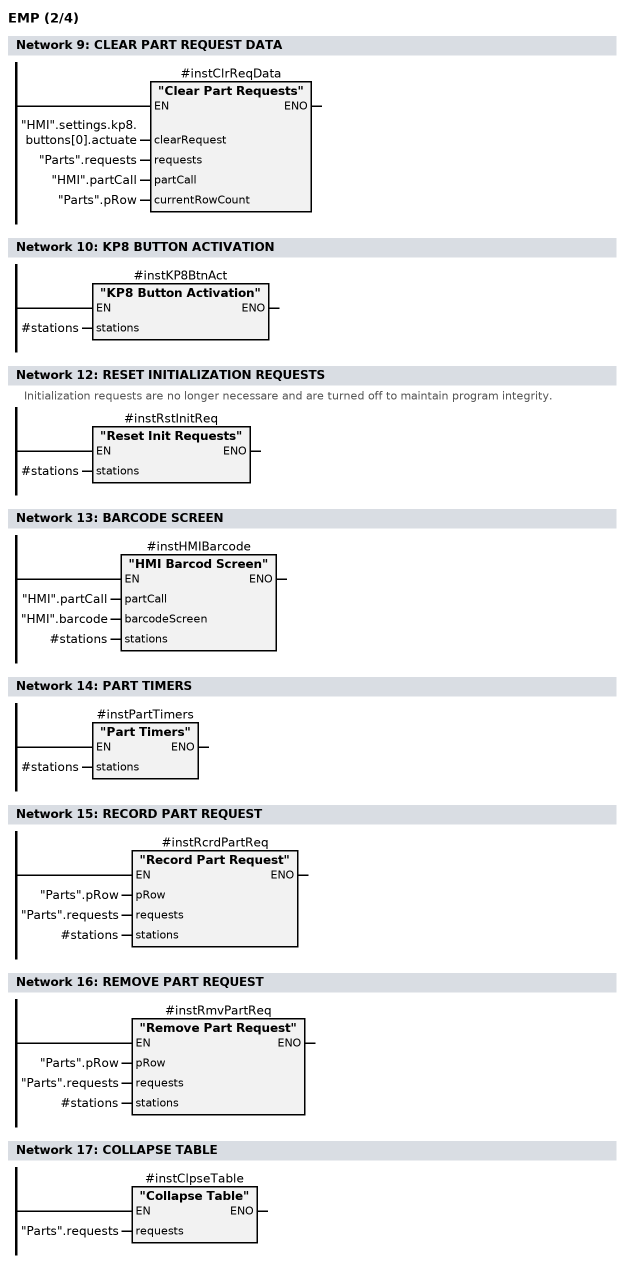
   RUNG wire#powerrail
      #instClrReqData(clearRequest := "HMI".settings.kp8.buttons[0].actuate, requests := "Parts".requests, partCall := "HMI".partCall, currentRowCount := "Parts".pRow)
   END_RUNG
   // the same network as SCL:
   #instClrReqData(clearRequest := "HMI".settings.kp8.buttons[0].actuate,   // "Clear Part Requests"
                   requests := "Parts".requests,
                   partCall := "HMI".partCall,
                   currentRowCount := "Parts".pRow);
END_REGION

REGION Network 10: KP8 BUTTON ACTIVATION
   RUNG wire#powerrail
      #instKP8BtnAct(stations := #stations)
   END_RUNG
   // the same network as SCL:
   #instKP8BtnAct(stations := #stations);   // "KP8 Button Activation"
END_REGION

REGION Network 11 (SCL): KP8 DRIVER CALLS
   REGION "LOOP THROUGH STATIONS"
       FOR #i := 0 TO "stnCount" DO
           #instKP8Drvs[#i](btnIn := #stations.me[#i].kp8In,
                            hardInit := #stations.me[#i].init.hard,
                            softInit := #stations.me[#i].init.soft,
                            btn0Activate := #stations.me[#i].kp8Config.activate[0],
                            btn0Mode := #stations.me[#i].kp8Config.mode[0],
                            btn0Group := #stations.me[#i].kp8Config.group[0],
                            btn0Flash := #stations.me[#i].kp8Config.flash[0],
                            btn0ColorOn1 := #stations.me[#i].kp8Config.colorOn1[0],
                            btn0ColorOn2 := #stations.me[#i].kp8Config.colorOn2[0],
                            btn0ColorOff := #stations.me[#i].kp8Config.colorOff[0],
                            btn1Activate := #stations.me[#i].kp8Config.activate[1],
                            btn1Mode := #stations.me[#i].kp8Config.mode[1],
                            btn1Group := #stations.me[#i].kp8Config.group[1],
                            btn1Flash := #stations.me[#i].kp8Config.flash[1],
                            btn1ColorOn1 := #stations.me[#i].kp8Config.colorOn1[1],
                            btn1ColorOn2 := #stations.me[#i].kp8Config.colorOn2[1],
                            btn1ColorOff := #stations.me[#i].kp8Config.colorOff[1],
                            btn2Activate := #stations.me[#i].kp8Config.activate[2],
                            btn2Mode := #stations.me[#i].kp8Config.mode[2],
                            btn2Group := #stations.me[#i].kp8Config.group[2],
                            btn2Flash := #stations.me[#i].kp8Config.flash[2],
                            btn2ColorOn1 := #stations.me[#i].kp8Config.colorOn1[2],
                            btn2ColorOn2 := #stations.me[#i].kp8Config.colorOn2[2],
                            btn2ColorOff := #stations.me[#i].kp8Config.colorOff[2],
                            btn3Activate := #stations.me[#i].kp8Config.activate[3],
                            btn3Mode := #stations.me[#i].kp8Config.mode[3],
                            btn3Group := #stations.me[#i].kp8Config.group[3],
                            btn3Flash := #stations.me[#i].kp8Config.flash[3],
                            btn3ColorOn1 := #stations.me[#i].kp8Config.colorOn1[3],
                            btn3ColorOn2 := #stations.me[#i].kp8Config.colorOn2[3],
                            btn3ColorOff := #stations.me[#i].kp8Config.colorOff[3],
                            btn4Activate := #stations.me[#i].kp8Config.activate[4],
                            btn4Mode := #stations.me[#i].kp8Config.mode[4],
                            btn4Group := #stations.me[#i].kp8Config.group[4],
                            btn4Flash := #stations.me[#i].kp8Config.flash[4],
                            btn4ColorOn1 := #stations.me[#i].kp8Config.colorOn1[4],
                            btn4ColorOn2 := #stations.me[#i].kp8Config.colorOn2[4],
                            btn4ColorOff := #stations.me[#i].kp8Config.colorOff[4],
                            btn5Activate := #stations.me[#i].kp8Config.activate[5],
                            btn5Mode := #stations.me[#i].kp8Config.mode[5],
                            btn5Group := #stations.me[#i].kp8Config.group[5],
                            btn5Flash := #stations.me[#i].kp8Config.flash[5],
                            btn5ColorOn1 := #stations.me[#i].kp8Config.colorOn1[5],
                            btn5ColorOn2 := #stations.me[#i].kp8Config.colorOn2[5],
                            btn5ColorOff := #stations.me[#i].kp8Config.colorOff[5],
                            btn6Activate := #stations.me[#i].kp8Config.activate[6],
                            btn6Mode := #stations.me[#i].kp8Config.mode[6],
                            btn6Group := #stations.me[#i].kp8Config.group[6],
                            btn6Flash := #stations.me[#i].kp8Config.flash[6],
                            btn6ColorOn1 := #stations.me[#i].kp8Config.colorOn1[6],
                            btn6ColorOn2 := #stations.me[#i].kp8Config.colorOn2[6],
                            btn6ColorOff := #stations.me[#i].kp8Config.colorOff[6],
                            btn7Activate := #stations.me[#i].kp8Config.activate[7],
                            btn7Mode := #stations.me[#i].kp8Config.mode[7],
                            btn7Group := #stations.me[#i].kp8Config.group[7],
                            btn7Flash := #stations.me[#i].kp8Config.flash[7],
                            btn7ColorOn1 := #stations.me[#i].kp8Config.colorOn1[7],
                            btn7ColorOn2 := #stations.me[#i].kp8Config.colorOn2[7],
                            btn7ColorOff := #stations.me[#i].kp8Config.colorOff[7],
                            btnStatesOut => #stations.me[#i].btnStates,
                            btnColorsOut => #stations.me[#i].kp8Out);
       END_FOR;
   END_REGION
END_REGION

REGION Network 12: RESET INITIALIZATION REQUESTS
   // Initialization requests are no longer necessare and are turned off to maintain program integrity.
   RUNG wire#powerrail
      #instRstInitReq(stations := #stations)
   END_RUNG
   // the same network as SCL:
   #instRstInitReq(stations := #stations);   // "Reset Init Requests"
END_REGION

REGION Network 13: BARCODE SCREEN
   RUNG wire#powerrail
      #instHMIBarcode(partCall := "HMI".partCall, barcodeScreen := "HMI".barcode, stations := #stations)
   END_RUNG
   // the same network as SCL:
   #instHMIBarcode(partCall := "HMI".partCall, barcodeScreen := "HMI".barcode, stations := #stations);   // "HMI Barcod Screen"
END_REGION

REGION Network 14: PART TIMERS
   RUNG wire#powerrail
      #instPartTimers(stations := #stations)
   END_RUNG
   // the same network as SCL:
   #instPartTimers(stations := #stations);   // "Part Timers"
END_REGION

REGION Network 15: RECORD PART REQUEST
   RUNG wire#powerrail
      #instRcrdPartReq(pRow := "Parts".pRow, requests := "Parts".requests, stations := #stations)
   END_RUNG
   // the same network as SCL:
   #instRcrdPartReq(pRow := "Parts".pRow, requests := "Parts".requests, stations := #stations);   // "Record Part Request"
END_REGION

REGION Network 16: REMOVE PART REQUEST
   RUNG wire#powerrail
      #instRmvPartReq(pRow := "Parts".pRow, requests := "Parts".requests, stations := #stations)
   END_RUNG
   // the same network as SCL:
   #instRmvPartReq(pRow := "Parts".pRow, requests := "Parts".requests, stations := #stations);   // "Remove Part Request"
END_REGION

REGION Network 17: COLLAPSE TABLE
   RUNG wire#powerrail
      #instClpseTable(requests := "Parts".requests)
   END_RUNG
   // the same network as SCL:
   #instClpseTable(requests := "Parts".requests);   // "Collapse Table"
END_REGION

REGION Network 18: LOG REQUESTS
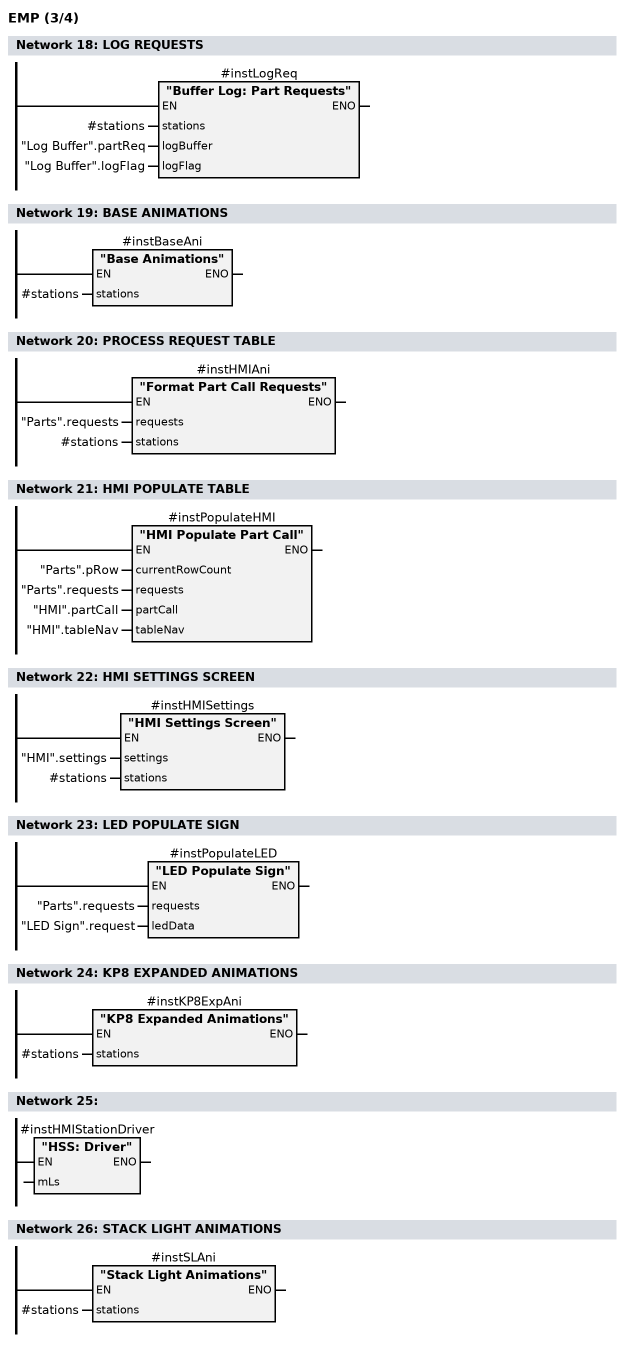
   RUNG wire#powerrail
      #instLogReq(stations := #stations, logBuffer := "Log Buffer".partReq, logFlag := "Log Buffer".logFlag)
   END_RUNG
   // the same network as SCL:
   #instLogReq(stations := #stations, logBuffer := "Log Buffer".partReq, logFlag := "Log Buffer".logFlag);   // "Buffer Log: Part Requests"
END_REGION

REGION Network 19: BASE ANIMATIONS
   RUNG wire#powerrail
      #instBaseAni(stations := #stations)
   END_RUNG
   // the same network as SCL:
   #instBaseAni(stations := #stations);   // "Base Animations"
END_REGION

REGION Network 20: PROCESS REQUEST TABLE
   RUNG wire#powerrail
      #instHMIAni(requests := "Parts".requests, stations := #stations)
   END_RUNG
   // the same network as SCL:
   #instHMIAni(requests := "Parts".requests, stations := #stations);   // "Format Part Call Requests"
END_REGION

REGION Network 21: HMI POPULATE TABLE
   RUNG wire#powerrail
      #instPopulateHMI(currentRowCount := "Parts".pRow, requests := "Parts".requests, partCall := "HMI".partCall, tableNav := "HMI".tableNav)
   END_RUNG
   // the same network as SCL:
   #instPopulateHMI(currentRowCount := "Parts".pRow,   // "HMI Populate Part Call"
                    requests := "Parts".requests,
                    partCall := "HMI".partCall,
                    tableNav := "HMI".tableNav);
END_REGION

REGION Network 22: HMI SETTINGS SCREEN
   RUNG wire#powerrail
      #instHMISettings(settings := "HMI".settings, stations := #stations)
   END_RUNG
   // the same network as SCL:
   #instHMISettings(settings := "HMI".settings, stations := #stations);   // "HMI Settings Screen"
END_REGION

REGION Network 23: LED POPULATE SIGN
   RUNG wire#powerrail
      #instPopulateLED(requests := "Parts".requests, ledData := "LED Sign".request)
   END_RUNG
   // the same network as SCL:
   #instPopulateLED(requests := "Parts".requests, ledData := "LED Sign".request);   // "LED Populate Sign"
END_REGION

REGION Network 24: KP8 EXPANDED ANIMATIONS
   RUNG wire#powerrail
      #instKP8ExpAni(stations := #stations)
   END_RUNG
   // the same network as SCL:
   #instKP8ExpAni(stations := #stations);   // "KP8 Expanded Animations"
END_REGION

REGION Network 25
   RUNG wire#powerrail
      #instHMIStationDriver(mLs :=)
   END_RUNG
   // the same network as SCL:
   #instHMIStationDriver();   // "HSS: Driver"
END_REGION

REGION Network 26: STACK LIGHT ANIMATIONS
   RUNG wire#powerrail
      #instSLAni(stations := #stations)
   END_RUNG
   // the same network as SCL:
   #instSLAni(stations := #stations);   // "Stack Light Animations"
END_REGION

REGION Network 27: GLOBAL TO SIMULATION
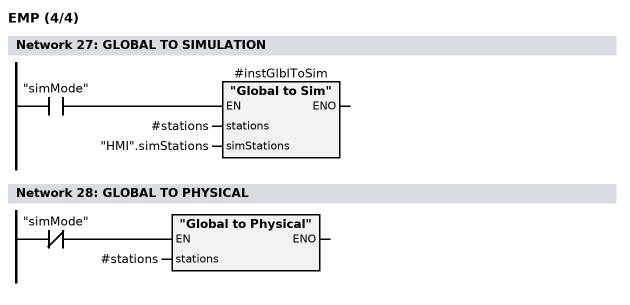
   RUNG wire#powerrail
      Contact( "simMode" )
      #instGlblToSim(stations := #stations, simStations := "HMI".simStations)
   END_RUNG
   // the same network as SCL:
   IF "simMode" THEN
       #instGlblToSim(stations := #stations, simStations := "HMI".simStations);   // "Global to Sim"
   END_IF;
END_REGION

REGION Network 28: GLOBAL TO PHYSICAL
   RUNG wire#powerrail
      I_Contact( "simMode" )
      "Global to Physical"(stations := #stations)
   END_RUNG
   // the same network as SCL:
   IF NOT "simMode" THEN "Global to Physical"(stations := #stations); END_IF;
END_REGION
END_FUNCTION_BLOCK

// folder: HMI Select Station

FUNCTION_BLOCK "HSS: Driver"   // FB32, LAD
{ S7_Optimized_Access := 'TRUE' }
VERSION : 0.1
   VAR_INPUT
      mLs : "Menu: Libraries";
   END_VAR
   VAR
      recipeSelector : Int;
      r1 : DInt;
      instHSSMenuSelection : "HSS: Menu Selection";
   END_VAR
   VAR_TEMP
      i : Int;
   END_VAR
BEGIN

REGION Network 1
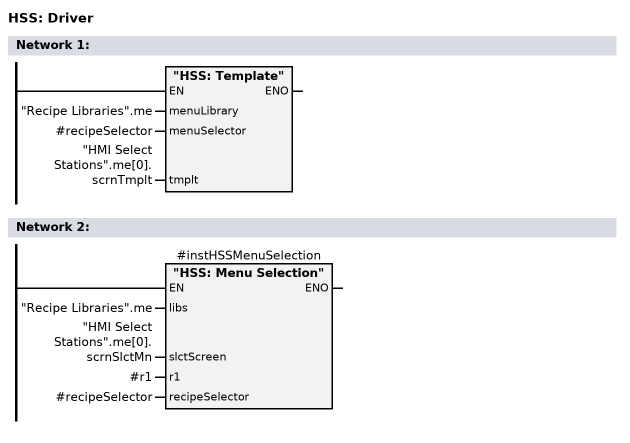
   RUNG wire#powerrail
      "HSS: Template"(menuLibrary := "Recipe Libraries".me, menuSelector := #recipeSelector, tmplt := "HMI Select Stations".me[0].scrnTmplt)
   END_RUNG
   // the same network as SCL:
   "HSS: Template"(menuLibrary := "Recipe Libraries".me,
                   menuSelector := #recipeSelector,
                   tmplt := "HMI Select Stations".me[0].scrnTmplt);
END_REGION

REGION Network 2
   RUNG wire#powerrail
      #instHSSMenuSelection(libs := "Recipe Libraries".me, slctScreen := "HMI Select Stations".me[0].scrnSlctMn, r1 := #r1, recipeSelector := #recipeSelector)
   END_RUNG
   // the same network as SCL:
   #instHSSMenuSelection(libs := "Recipe Libraries".me,   // "HSS: Menu Selection"
                         slctScreen := "HMI Select Stations".me[0].scrnSlctMn,
                         r1 := #r1,
                         recipeSelector := #recipeSelector);
END_REGION
END_FUNCTION_BLOCK

FUNCTION_BLOCK "HSS: Part Selection"   // FB33, SCL
{ S7_Optimized_Access := 'TRUE' }
VERSION : 0.1
BEGIN
END_FUNCTION_BLOCK

FUNCTION_BLOCK "HSS: Menu Selection"   // FB35, SCL
{ S7_Optimized_Access := 'TRUE' }
VERSION : 0.1
   VAR_INPUT
      libs : "Menu: Libraries";
   END_VAR
   VAR_IN_OUT
      slctScreen : "HSS: Menu Selection Screen";
      r1 : DInt;
      recipeSelector : Int;
   END_VAR
   VAR
      old : Struct
         navPress : Bool;
      END_STRUCT;
      instTableNavigation : "Table Navigatio";
   END_VAR
   VAR_TEMP
      eval : "HSS: Menu Selection Screen";
      pbs : Array[0..#pbFlagCnt] of Bool;
      POS : DInt;
      status : DInt;
      i : Int;
      btnNum : Int;
      pRowVisLbl : Int;
      pRowInvisLbl : Int;
      pRecipeInvisLbl : Int;
      pRecipeVisLbl : Int;
      pRecipeLib : Int;
      pRowTxt : Int;
      pRecipeTxt : Int;
      shifter : DWord;
      btnsAsBool : Array[0..31] of Bool;
      rows : Array[0..99] of DInt;
      offset : DInt;
      navPress : Bool;
      selPress : Bool;
      maxRows : DInt;
   END_VAR
   VAR CONSTANT
      pbFlagCnt : Int := 31;
      btnCnt : Int := 5;
      navMask : DWord := 16#0000_003F;
      visRows : DInt := 6;
      home : DInt := -1000;
      end : DInt := -2000;
   END_VAR
BEGIN
   REGION "INITITALIZE LOCALS"
       #eval := #slctScreen;
       #maxRows := #libs.stations[24].size;
       SCATTER(IN := #eval.pbs,
               OUT => #btnsAsBool);
   END_REGION


   REGION "GET RECIPE SELECTION PRESS" 
       FOR #i := 6 TO 31 DO
           IF #btnsAsBool[#i] THEN
               #recipeSelector := DINT_TO_INT(#r1) + #i - 6;
               #selPress := TRUE;
               EXIT;
           END_IF;
       END_FOR;
   END_REGION


   REGION "TABLE NAVIGATION"
       IF "HMI Select Stations".me[0].scrnSlctMn.pbs.%X0 THEN
           #offset := #home;
       END_IF;
       IF "HMI Select Stations".me[0].scrnSlctMn.pbs.%X1 THEN
           #offset := -1 * #visRows;
       END_IF;
       IF "HMI Select Stations".me[0].scrnSlctMn.pbs.%X2 THEN
           #offset := -1;
       END_IF;
       IF "HMI Select Stations".me[0].scrnSlctMn.pbs.%X3 THEN
           #offset := 1;
       END_IF;
       IF "HMI Select Stations".me[0].scrnSlctMn.pbs.%X4 THEN
           #offset := #visRows;
       END_IF;
       IF "HMI Select Stations".me[0].scrnSlctMn.pbs.%X5 THEN
           #offset := #end;
       END_IF;

       IF ("HMI Select Stations".me[0].scrnSlctMn.pbs AND #navMask) <> 0 THEN
           #navPress := true;
       END_IF;

       #instTableNavigation(maxRows := #maxRows,
                            visRows := #visRows,
                            offset := #offset,
                            trigger := #navPress,
                            r1 := #r1,
                            rowIndices := #rows);
   END_REGION


   REGION "LABELS"
       IF #navPress AND NOT #old.navPress THEN
           FOR #i := 0 TO #visRows - 1 DO
               "Recipe Nav Button"(visRows := DINT_TO_INT(#visRows),
                                   actuate := #btnsAsBool[#i],
                                   maxRows := DINT_TO_INT(#maxRows),
                                   btnNum := #i,
                                   recipeSelectScreen := #eval);
               "Recipe Select Button"(visRows := DINT_TO_INT(#visRows),
                                      rowNum := DINT_TO_INT(#rows[#i]),
                                      lib := #libs.stations[24],
                                      actuate := #btnsAsBool[#i + 6],
                                      maxRows := DINT_TO_INT(#maxRows),
                                      btnNum := #i,
                                      recipeSelectScreen := #eval);
           END_FOR;
       END_IF;
   END_REGION


   REGION "CHANGE DETECTION"
       #old.navPress := #navPress;
   END_REGION


   REGION "COPY TO GLOBAL"
       #slctScreen := #eval;
   END_REGION
END_FUNCTION_BLOCK

FUNCTION "HSS: Template" : Void   // FC24, SCL
{ S7_Optimized_Access := 'TRUE' }
VERSION : 0.1
   VAR_INPUT
      menuLibrary : "Menu: Libraries";
      menuSelector : Int;
   END_VAR
   VAR_IN_OUT
      tmplt : "HSS: Template Screen";
   END_VAR
   VAR_TEMP
      i : Int;
   END_VAR
BEGIN
   #tmplt.animate[0] := "BgGray";
   #tmplt.text[0] := "Word Wrap"(stringIn := #menuLibrary.stations[24].entry[#menuSelector],
                                 maxLength := 26);
END_FUNCTION

// folder: Network Diagnostics

FUNCTION_BLOCK "NetDiag: Get IPs"   // FB27, SCL
{ S7_Optimized_Access := 'TRUE' }
VERSION : 0.1
   VAR_OUTPUT
      error : Bool := FALSE;   // Rising edge informs that an error occurred during the execution of the FB
      status : Word := 16#0000;   // Current status of FB
      statusID : Word := 16#0;   // Current status ID of calling instruction
   END_VAR
   VAR_IN_OUT
      ioSystemData : "UserDiag_typeIOSystem";   // IO-System diagnostics data
   END_VAR
   VAR
      statError : Bool := FALSE;   // Static value for output error
      statStatus : Word := 16#0000;   // Static value for output status
      statStatusID : Word := 16#0;   // Static value for output statusID
      instGetStationInfo : GetStationInfo;   // Instance of GetStationInfo
      statFirstDeviceFlag : Bool := TRUE;   // Help tag for the first device in the linked list
      statDeviceIndex : Int := 0;   // Device/slave index
   END_VAR
   VAR_TEMP
      tempIP : IF_CONF_v4;   // Temporary IP address
   END_VAR
   VAR CONSTANT
      STATUS_EXECUTION_FINISHED : Word := 16#0000;   // Execution finished without errors
      ID_GET_STATION_INFO : Word := 12;   // StatusID during GetStationInfo command
      MODE_IPV4 : UInt := 1;   // Address parameter according to IPv4
      LAST_DEVICE : Int := -1;   // No next device
   END_VAR
BEGIN
   //=============================================================================
   //SIEMENS AG
   //(c)Copyright 2015 All Rights Reserved
   //-----------------------------------------------------------------------------
   //Library: 
   //Tested with: S7-1516-3 PN/DP FW 2.5
   //Engineering: TIA Portal V15
   //Restrictions: Call in cyclic OB
   //Requirements: -
   //Functionality: Get IP address of IO devices
   //-----------------------------------------------------------------------------
   //Change log table:
   //Version  Date       Expert in charge                Changes applied
   //01.00.00 20.12.2017 Siemens Industry Online Support First released version
   //=============================================================================

   //=============================================================================
   // Go through existing devices and get IP address
   //=============================================================================
   // Initialize the pointer for the first run 
   IF (#statFirstDeviceFlag = TRUE)
   THEN
       #statDeviceIndex := #ioSystemData.firstDevice;
       #statFirstDeviceFlag := FALSE;
   END_IF;

   // Check and store the IP address, if the device is existing
   // GetStationInfo is an acyclic instruction. In the FB, the
   // instruction has to be repeated until it is done or error
   IF ((#ioSystemData.number >= 100)
       AND (#ioSystemData.number <= 115)
       AND (#ioSystemData.devices[#statDeviceIndex].exists = TRUE)
       AND (#ioSystemData.devices[#statDeviceIndex].ipAddress.ADDR[1] = 0))
   THEN
       // Get IP address of each decive in PN System
       #instGetStationInfo(REQ := TRUE,
                           LADDR := #ioSystemData.devices[#statDeviceIndex].hardwareId,
                           MODE := #MODE_IPV4,
                           DATA := #tempIP);

       IF (#instGetStationInfo.ERROR = TRUE)
       THEN
           // Error handling
           #statStatus := #instGetStationInfo.STATUS;
           #statStatusID := #ID_GET_STATION_INFO;
           #statError := TRUE;

           // Everything is ok --> Copy IP address    
       ELSIF (#instGetStationInfo.DONE = TRUE)
       THEN
           #ioSystemData.devices[#statDeviceIndex].ipAddress := #tempIP.InterfaceAddress;

           // Initialize the pointer for the next run
           #statDeviceIndex := #ioSystemData.devices[#statDeviceIndex].nextDevice;
       ELSE
           ;
       END_IF;
   ELSE
       // Initialize the pointer for the next run
       #statDeviceIndex := #ioSystemData.devices[#statDeviceIndex].nextDevice;
   END_IF;

   // Check last device
   IF (#statDeviceIndex = #LAST_DEVICE)
   THEN
       #statDeviceIndex := #ioSystemData.firstDevice;
   END_IF;

   // Write static values to outputs
   #error := #statError;
   #status := #statStatus;
   #statusID := #statStatusID;
END_FUNCTION_BLOCK

FUNCTION_BLOCK "NetDiag: Coordinate"   // FB28, LAD
{ S7_Optimized_Access := 'TRUE' }
VERSION : 0.1
// //============================================================================
// //SIEMENS AG
// //(c)Copyright 2017 All Rights Reserved
// //-----------------------------------------------------------------------------
// //Library: -
// //Tested with: S7-1516-3 PN/DP FW 2.5
// //Engineering: TIA Portal V15
// //Restrictions: -
// //Requirements: -
// //Functionality: Main FB for diagnostics
// //-----------------------------------------------------------------------------
// //Change log table:
// //Version  Date              Expert in charge                               Changes applied
// //01.00.00 25.04.2017 Siemens Industry Online Support First released version
// //01.01.00 01.12.2017 Siemens Industry Online Support Renamed in "UserDiag_Diagnostics"
// //                                                                                                    Check Flag "startDiag"
// //============================================================================
   VAR_IN_OUT
      startDiag : Bool := false;   // Startflag for diagnostic
      plcData : "UserDiag_typePLC";   // PLC diagnostics data
      ioSystemData : Array[1.."USERDIAG_IO_SYSTEMS_UPPER_LIM"] of "UserDiag_typeIOSystem";   // IO-System diagnostics data
   END_VAR
   VAR
      instPLCChk : "NetDiag: Check PLC";   // Instance of "UserDiag_PLCCheck"
      instIOSysChk : "NetDiag: IO Systems";   // Instance of "UserDiag_IOSystemCheck"
   END_VAR
BEGIN

REGION Network 1: Check Startflag for diagnostic
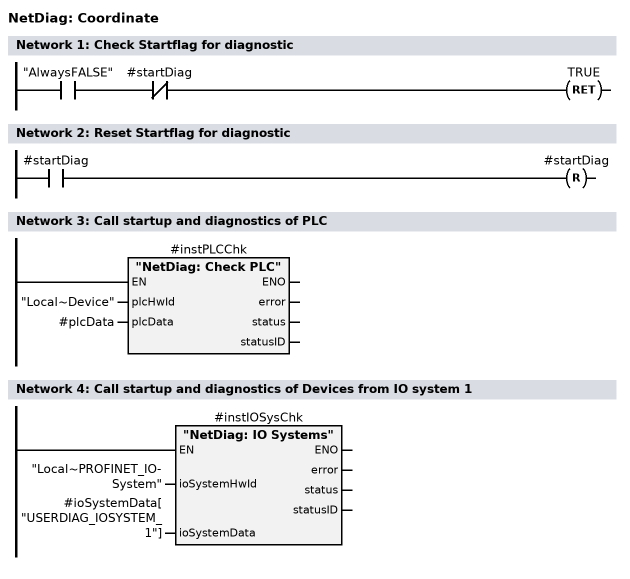
   IF "AlwaysFALSE" AND NOT #startDiag THEN
       ENO := TRUE;
       RETURN;
   END_IF;
END_REGION

REGION Network 2: Reset Startflag for diagnostic
   RUNG wire#powerrail
      Contact( #startDiag )
      R_Coil( #startDiag )
   END_RUNG
   // the same network as SCL:
   IF #startDiag THEN #startDiag := FALSE; END_IF;
END_REGION

REGION Network 3: Call startup and diagnostics of PLC
   RUNG wire#powerrail
      #instPLCChk(plcHwId := "Local~Device", plcData := #plcData, error =>, status =>, statusID =>)
   END_RUNG
   // the same network as SCL:
   #instPLCChk(plcHwId := "Local~Device", plcData := #plcData);   // "NetDiag: Check PLC"
END_REGION

REGION Network 4: Call startup and diagnostics of Devices from IO system 1
   RUNG wire#powerrail
      #instIOSysChk(ioSystemHwId := "Local~PROFINET_IO-System", ioSystemData := #ioSystemData["USERDIAG_IOSYSTEM_1"], error =>, status =>, statusID =>)
   END_RUNG
   // the same network as SCL:
   #instIOSysChk(ioSystemHwId := "Local~PROFINET_IO-System",   // "NetDiag: IO Systems"
                 ioSystemData := #ioSystemData["USERDIAG_IOSYSTEM_1"]);
END_REGION
END_FUNCTION_BLOCK

FUNCTION_BLOCK "NetDiag: Check PLC"   // FB29, SCL
{ S7_Optimized_Access := 'TRUE' }
VERSION : 0.1
   VAR_INPUT
      plcHwId : Hw_Device := 0;   // Hardware ID
   END_VAR
   VAR_OUTPUT
      error : Bool := FALSE;   // Rising edge informs that an error occurred during the execution of the FB
      status : Word := 16#0000;   // Current status of FB
      statusID : Word := 16#0;   // Current status ID of calling instruction
   END_VAR
   VAR_IN_OUT
      plcData : "UserDiag_typePLC";   // PLC diagnostics data
   END_VAR
   VAR
      statError : Bool := FALSE;   // Static value for output error
      statStatus : Word := 16#0000;   // Static value for output status
      statStatusID : Word := 16#0;   // Static value for output statusID
      statGeoAddr : GEOADDR;   // Slot information
      statGeoLaddr : Hw_Any := 16#0000;   // GEO2LOG hardware identifier
      statProblemPlcModulStates : Array[0..#MODULES_STATES_UPPER_LIM] of Bool;   // Storage of the status of all modules in the PLC central station --> State: Problem
      statFaultyPlcModulStates : Array[0..#MODULES_STATES_UPPER_LIM] of Bool;   // Storage of the status of all modules in the PLC central station --> State: Faulty
      statExistingPlcModulStates : Array[0..#MODULES_STATES_UPPER_LIM] of Bool;   // Storage of the status of all modules in the PLC central station --> State: Exists
      statActualCentralModules : USInt := 0;   // Actual number of modules in the central station (PLC)
   END_VAR
   VAR_TEMP
      tempSlotNum : Int;   // Index slot number
      tempRetValGeo : Int;   // GEO2LOG error information
      tempRetValModuleStates : Int;   // Return value system function ModuleStates
   END_VAR
   VAR CONSTANT
      STATUS_EXECUTION_FINISHED : Word := 16#0000;   // Execution finished without errors
      ERR_MAX_SLOTS_PER_PLC : Word := 16#8400;   // There are more modules configured as defined with the user constant: USERDIAG_SLOTS_PER_PLC_UPPER_LIM
      ID_LOCAL : Word := 1;   // StatusID local
      ID_MODULE_STATES_CONFIGURED : Word := 2;   // StatusID during ModuleStates command (configured mode)
      ID_MODULE_STATES_FAULTY : Word := 3;   // StatusID during ModuleStates command (faulty mode)
      ID_MODULE_STATES_PROBLEM : Word := 4;   // StatusID during ModuleStates command (problem mode)
      ID_MODULE_STATES_EXISTING : Word := 5;   // StatusID during ModuleStates command (existing mode)
      ID_LED : Word := 12;   // StatusID occurred during LED command
      MODE_FAULTY : USInt := 2;   // Used for instruction DeviceStates, read out all faulty devices
      MODE_EXIST : USInt := 4;   // Used for instruction DeviceStates, read out all devices not reachable
      MODE_PROBLEM : USInt := 5;   // Used for instruction DeviceStates, read out all devices with several problems
      STATE_OK : USInt := 1;   // Module state: ok
      STATE_FAULT : USInt := 2;   // Modulestate: fault
      STATE_PROBLEM : USInt := 5;   // Module state: problem
      STATE_WAS_FAULT : USInt := 12;   // Module state: was fault
      STATE_PROBLEM_GONE : USInt := 15;   // Module state: had a problem
      MODULE_OF_PLC : USInt := 4;   // GEO2LOG structure: HW type = 4
      CPU : USInt := 0;   // GEO2LOG structure: Area = 0
      CENTRAL_SYSTEM : USInt := 0;   // GEO2LOG structure: IO System = 0
      CENTRAL_STATION : USInt := 0;   // GEO2LOG structure: Station = 0
      NO_LED : Int := 0;   // LED does not exist
      LED_OFF : Int := 1;   // LED is permanently switched off
      LED_NO_INFO : Int := 9;   // LED exists, but status information not available
      MODULES_STATES_UPPER_LIM : Int := 127;   // Upper array limit for output tag of instruction ModuleStates
      ERROR_LED : UInt := 2;   // Identification number of the LED
   END_VAR
BEGIN
   //=============================================================================
   //SIEMENS AG
   //(c)Copyright 2017 All Rights Reserved
   //-----------------------------------------------------------------------------
   //Library: 
   //Tested with: S7-1516-3 PN/DP FW 2.5
   //Engineering: TIA Portal V15
   //Restrictions: Call in cyclic OB
   //Requirements: -
   //Functionality: Determine plc state and local module states
   //-----------------------------------------------------------------------------
   //Change log table:
   //Version  Date       Expert in charge                Changes applied
   //01.00.00 27.01.2017 Siemens Industry Online Support First released version
   //01.00.01 20.12.2017 Siemens Industry Online Support actualConfiguredSlots >= 1
   //01.00.02 27.02.2018 Siemens Industry Online Support Minor corrections
   //=============================================================================

   IF (#plcData.hardwareId = 0)
   THEN
       #statGeoAddr.HWTYPE := #MODULE_OF_PLC;      // Hardware type 4: module
       #statGeoAddr.AREA := #CPU;                  // Area ID 0: CPU
       #statGeoAddr.IOSYSTEM := #CENTRAL_SYSTEM;   // PROFINET IO system (0 = central unit in the rack)
       #statGeoAddr.STATION := #CENTRAL_STATION;   // Number of the rack if area identifier AREA = 0 (central module)

       #statStatus := #STATUS_EXECUTION_FINISHED;
       #statStatusID := 0;
       #statError := FALSE;
       #statActualCentralModules := 0;

       FOR #tempSlotNum := 0 TO "USERDIAG_SLOTS_PER_PLC_UPPER_LIM" DO
           // Slot number
           #statGeoAddr.SLOT := INT_TO_UINT(#tempSlotNum);
           // read LADDR from local modules
           #tempRetValGeo := GEO2LOG(GEOADDR := #statGeoAddr,
                                     LADDR => #statGeoLaddr);
           // Check Retval
           IF ((#tempRetValGeo = 0)
               AND (#statGeoLaddr <> 16#0))
           THEN
               // Store LADDR from local modules in diagnostic data block
               IF (#tempSlotNum = 1)
               THEN
                   #plcData.hardwareId := #statGeoLaddr;
               END_IF;
               #plcData.slots[#tempSlotNum].hardwareId := #statGeoLaddr;
               #statActualCentralModules := #statActualCentralModules + 1;
               #plcData.slots[#tempSlotNum].configured := TRUE;
           ELSE
               // If the return value ist not = 0 --> the device/system/module is not
               // configured --> No error handling
               // set LADDR from local modules to 0 in diagnostic data block
               #plcData.slots[#tempSlotNum].hardwareId := 0;
               #plcData.slots[#tempSlotNum].configured := FALSE;
           END_IF;
           // Store the actual configured devices in the diagnostics DB
           #plcData.actualConfiguredSlots := #statActualCentralModules;
       END_FOR;

       // Check if further slots are configured
       #statGeoAddr.SLOT := INT_TO_UINT(#tempSlotNum);

       #tempRetValGeo := GEO2LOG(GEOADDR := #statGeoAddr,
                                 LADDR => #statGeoLaddr);

       IF ((#tempRetValGeo = 0)
           AND (#statGeoLaddr <> 16#0))
       THEN
           // In the PLC are more slots configured as defined with the user constant
           #statStatus := #ERR_MAX_SLOTS_PER_PLC;
           #statStatusID := #ID_LOCAL;
           #statError := TRUE;
       END_IF;

   END_IF;

   // Reset PLC error state
   #plcData.error := FALSE;

   //=============================================================================
   // Check modul states from LOCAL MODULES
   //=============================================================================
   // Check if central module are available - at least one module is always
   // configured, the PLC itself
   IF (#plcData.actualConfiguredSlots >= 1)
   THEN

       // Check the status of the local modules
       #tempRetValModuleStates := ModuleStates(LADDR := #plcHwId,
                                               MODE := #MODE_PROBLEM,
                                               STATE := #statProblemPlcModulStates);

       // Check if the block call was successful
       IF (#tempRetValModuleStates <> 0)
       THEN
           // Error handling
           #statStatus := INT_TO_WORD(#tempRetValModuleStates);
           #statStatusID := #ID_MODULE_STATES_PROBLEM;
           #statError := TRUE;
       ELSE
           ; // Everything is ok!
       END_IF;

       #tempRetValModuleStates := ModuleStates(LADDR := #plcHwId,
                                               MODE := #MODE_FAULTY,
                                               STATE := #statFaultyPlcModulStates);

       // Check if the block call was successful
       IF (#tempRetValModuleStates <> 0)
       THEN
           // Error handling
           #statStatus := INT_TO_WORD(#tempRetValModuleStates);
           #statStatusID := #ID_MODULE_STATES_FAULTY;
           #statError := TRUE;
       ELSE
           ; // Everything is ok!
       END_IF;

       #tempRetValModuleStates := ModuleStates(LADDR := #plcHwId,
                                               MODE := #MODE_EXIST,
                                               STATE := #statExistingPlcModulStates);

       // Check if the block call was successful
       IF (#tempRetValModuleStates <> 0)
       THEN
           // Error handling
           #statStatus := INT_TO_WORD(#tempRetValModuleStates);
           #statStatusID := #ID_MODULE_STATES_EXISTING;
           #statError := TRUE;
       ELSE
           ; // Everything is ok!
       END_IF;

   ELSE
       ; // There are no central moduls configured
   END_IF;

   //=============================================================================
   // Set module states of LOCAL MODULES
   //=============================================================================
   #tempSlotNum := 0;
   WHILE (#tempSlotNum <= #plcData.actualConfiguredSlots)
   DO
       IF (#plcData.slots[#tempSlotNum].configured)
       THEN
           IF (#statExistingPlcModulStates[#tempSlotNum + 1] = TRUE)
           THEN
               #plcData.slots[#tempSlotNum].exists := TRUE;
               CASE #plcData.slots[#tempSlotNum].state OF
                   #STATE_WAS_FAULT,
                   #STATE_PROBLEM_GONE:
                       ;
                   #STATE_FAULT:
                       #plcData.slots[#tempSlotNum].state := #STATE_WAS_FAULT;
                   #STATE_PROBLEM:
                       #plcData.slots[#tempSlotNum].state := #STATE_PROBLEM_GONE;
                   ELSE
                       #plcData.slots[#tempSlotNum].state := #STATE_OK;
               END_CASE;
           ELSE
               #plcData.slots[#tempSlotNum].error := TRUE;
               #plcData.error := TRUE;
               #plcData.slots[#tempSlotNum].exists := FALSE;
           END_IF;

           IF (#statFaultyPlcModulStates[#tempSlotNum + 1] = TRUE)
           THEN
               // Modul is faulty
               #plcData.slots[#tempSlotNum].faulty := TRUE;
               #plcData.slots[#tempSlotNum].problem := TRUE;
               #plcData.slots[#tempSlotNum].error := TRUE;
               #plcData.slots[#tempSlotNum].state := #STATE_FAULT;
           ELSIF (#statProblemPlcModulStates[#tempSlotNum + 1] = TRUE)
           THEN
               // Modul has a problem
               #plcData.slots[#tempSlotNum].faulty := FALSE;
               #plcData.slots[#tempSlotNum].problem := TRUE;
               #plcData.slots[#tempSlotNum].error := TRUE;
               #plcData.slots[#tempSlotNum].state := #STATE_PROBLEM;
           ELSE
               // Modul is OK
               #plcData.slots[#tempSlotNum].error := FALSE;
               #plcData.slots[#tempSlotNum].problem := FALSE;
               #plcData.slots[#tempSlotNum].faulty := FALSE;
           END_IF;

           // Error in PLC - Slot = 1, but index must be increased by 1, because of bit 0 = group display
           // --> used index = 2
           IF (#statProblemPlcModulStates[2] = TRUE)
               OR (#statFaultyPlcModulStates[2] = TRUE)
           THEN
               #plcData.error := TRUE;
           END_IF;
       END_IF;

       #tempSlotNum := #tempSlotNum + 1;
   END_WHILE;

   // Write static values to outputs
   #error := #statError;
   #status := #statStatus;
   #statusID := #statStatusID;

   //----------------------------------------------------------------------------------------------
END_FUNCTION_BLOCK

FUNCTION_BLOCK "NetDiag: IO Systems"   // FB30, SCL
{ S7_Optimized_Access := 'TRUE' }
VERSION : 0.1
   VAR_INPUT
      ioSystemHwId : Hw_IoSystem := 16#0000;   // This ID is representing the IO System (PN or DP), find the ID in the system constants
   END_VAR
   VAR_OUTPUT
      error : Bool := FALSE;   // Rising edge informs that an error occurred during the execution of the FB
      status : Word := 16#0000;   // Current status of FB
      statusID : Word := 16#0;   // Current status ID of calling instruction
   END_VAR
   VAR_IN_OUT
      ioSystemData : "UserDiag_typeIOSystem";   // IO-System diagnostics data
   END_VAR
   VAR
      statError : Bool := FALSE;   // Static value for output error
      statStatus : Word := 16#0000;   // Static value for output status
      statStatusID : Word := 16#0;   // Static value for output statusID
      statActualConfiguredDevices : Int := 0;   // Actual number of devices/slaves in the IOSystem/DP-Mastersystem
      statGeoAddr : GEOADDR;   // Slot information
      statGeoLaddr : Hw_Any := 16#0000;   // GEO2LOG hardware identifier
      statConfiguredDevices : Array[0..#DEVICES_STATES_UPPER_LIM] of Bool;   // Temporary storage of the return of "DeviceStates", to combine the states of the devices/slaves with numbers and names
      statExistingDevices : Array[0..#DEVICES_STATES_UPPER_LIM] of Bool;   // Temporary storage of the return of "DeviceStates", to combine the states of the devices/slaves with numbers and names
      statFaultyDevices : Array[0..#DEVICES_STATES_UPPER_LIM] of Bool;   // Temporary storage of the return of "DeviceStates", to combine the states of the devices/slaves with numbers and names
      statDisabledDevices : Array[0..#DEVICES_STATES_UPPER_LIM] of Bool;   // Temporary storage of the return of "DeviceStates", to combine the states of the devices/slaves with numbers and names
      statProblemDevices : Array[0..#DEVICES_STATES_UPPER_LIM] of Bool;   // Temporary storage of the return of "DeviceStates", to combine the states of the devices/slaves with numbers and names
      statDeviceProblemModules : Array[0..#MODULES_STATES_UPPER_LIM] of Bool;   // Storage of the status of all modules in the PN Devices / PB Slaves --> State: Problem
      statDeviceFaultyModules : Array[0..#MODULES_STATES_UPPER_LIM] of Bool;   // Storage of the status of all modules in the PN Devices / PB Slaves --> State: Faulty
      statDeviceExistingModules : Array[0..#MODULES_STATES_UPPER_LIM] of Bool;   // Storage of the status of all modules in the PN Devices / PB Slaves --> State: Existing
      instGetNameDevices : Get_Name;   // Instance of the system function "GetName"
      statInitString : String := '';   // Used to initialize the temporary string to convert into STRING[50]
      statFirstDevice : UInt := 0;   // Station number of the first device of the list
      statFirstDeviceFlag : Bool := TRUE;   // Help tag for the first device in the linked list
      statLastDevice : UInt := 0;   // Station number of the last device of the list
      statMaxDevices : Int := 0;   // Max devices per IO system
   END_VAR
   VAR_TEMP
      tempIndex : Int;   // Index of configured devices/slaves
      tempDeviceIndex : Int;   // Device/slave index
      tempSlotIndex : Int;   // Slot index
      tempSlotNum : Int;   // Index module number
      tempRetValGeo : Int;   // GEO2LOG error information
      tempRetValDeviceStates : Int;   // DeviceStates error information
      tempRetValModuleStates : Int;   // Return value of the system function "ModuleStates"
      tempStringConvert : String;   // Store the device names temporary here, to convert them into STRING[50]
      tempLastDevice : UInt;   // Temporary storage of the actual index, if it´s the last device --> store it in static
      tempDeviceInit : "UserDiag_typeDevice";   // Initalization of the device/slave diagnostic structure
   END_VAR
   VAR CONSTANT
      STATUS_EXECUTION_FINISHED : Word := 16#0000;   // Execution finished without errors
      ERR_MAX_SLOTS_PER_DEVICE : Word := 16#8400;   // There are more modules configured as defined with the user constant: USERDIAG_SLOTS_PER_DEVICE_UPPER_LIM
      ERR_MAX_DEVICES_PER_IOSYSTEM : Word := 16#8401;   // There are more modules configured as defined with the user constant: USERDIAG_DEVICES_PER_IO_SYTEM_UPPER_LIM
      ID_LOCAL : Word := 1;   // StatusID local
      ID_MODULE_STATES_CONFIGURED : Word := 2;   // StatusID during ModuleStates command (configured mode)
      ID_MODULE_STATES_FAULTY : Word := 3;   // StatusID during ModuleStates command (faulty mode)
      ID_MODULE_STATES_PROBLEM : Word := 4;   // StatusID during ModuleStates command (problem mode)
      ID_MODULE_STATES_EXISTING : Word := 5;   // StatusID during ModuleStates command (existing mode)
      ID_DEVICE_STATES_CONFIGURED : Word := 6;   // StatusID during DeviceStates command (configuration mode)
      ID_DEVICE_STATES_FAULTY : Word := 7;   // StatusID during DeviceStates command (fault mode)
      ID_DEVICE_STATES_PROBLEM : Word := 8;   // StatusID during DeviceStates command (problem mode)
      ID_DEVICE_STATES_EXISTING : Word := 9;   // StatusID during DeviceStates command (existing mode)
      ID_DEVICE_STATES_DISABLED : Word := 10;   // StatusID during DeviceStates command (disable mode)
      ID_GET_NAME : Word := 11;   // StatusID during GET_NAME command
      MODE_CONFIGURED : USInt := 1;   // Used for instruction DeviceStates/ModuleStates, read out all configured devices/slaves
      MODE_FAULTY : USInt := 2;   // Used for instruction DeviceStates/ModuleStates, read out all faulty devices/slaves
      MODE_DISABLED : USInt := 3;   // Used for instruction DeviceStates/ModuleStates, read out all disabled devices/slaves
      MODE_EXIST : USInt := 4;   // Used for instruction DeviceStates/ModuleStates, read out all devices/slaves not reachable
      MODE_PROBLEM : USInt := 5;   // Used for instruction DeviceStates/ModuleStates, read out all devices with several problems
      DEVICE_SLAVE : USInt := 2;   // GEO2LOG structure: HW type = 2
      MODULE_OF_DEVICE : USInt := 4;   // GEO2LOG structure: HW type = 4
      IO_SYSTEM_AREA : USInt := 1;   // GEO2LOG structure: Area = 1
      DP_SYSTEM_AREA : USInt := 2;   // GEO2LOG structure: Area = 2
      STATE_OK : USInt := 1;   // Device/modul state: ok
      STATE_FAULT : USInt := 2;   // Device/modul state: fault
      STATE_LOST_CON : USInt := 3;   // Device/modul state: lost connection
      STATE_DISABLED : USInt := 4;   // Device/modul state: disabled
      STATE_PROBLEM : USInt := 5;   // Device/modul state: problem
      STATE_WAS_FAULT : USInt := 12;   // Device/modul state: was fault
      STATE_WAS_LOST : USInt := 13;   // Device/modul state: connection was lost
      STATE_WAS_DISABLED : USInt := 14;   // Device/modul state: device/slave was disabled
      STATE_PROBLEM_GONE : USInt := 15;   // Device/modul state: had a problem
      MODULES_STATES_UPPER_LIM : Int := 127;   // Upper array limit for output tag of instruction ModuleStates
      DEVICES_STATES_UPPER_LIM : Int := 1023;   // Upper array limit for output tag of instruction DeviceStates
      ERR_HWID_NOT_EXISTENT : Int := 16#8091;   // Hardware identifier of the LADDR parameter does not exist. Check (for example, in the system constants) whether the value for LADDR exists in the project.
      ERR_LADDR_ADDRESS : Int := 16#8092;   // LADDR does not address a PROFINET IO or DP master system.
      POS_FIRST_CHAR : Int := 50;   // Position of first character to be deleted
      NUMBER_CHAR : Int := 204;   // Number of characters to be deleted
      MAX_SLAVES_DP : Int := 127;   // Max number of slaves in a PROFIBUS IO system
      LAST_DEVICE : Int := -1;   // No next device
   END_VAR
BEGIN
   //=============================================================================
   //SIEMENS AG
   //(c)Copyright 2015 All Rights Reserved
   //-----------------------------------------------------------------------------
   //Library: 
   //Tested with: S7-1516-3 PN/DP FW 2.5
   //Engineering: TIA Portal V15
   //Restrictions: Call in cyclic OB
   //Requirements: -
   //Functionality: Determine hardware identifier and module states from local and
   //               device modules 
   //-----------------------------------------------------------------------------
   //Change log table:
   //Version  Date       Expert in charge                Changes applied
   //01.00.00 27.01.2017 Siemens Industry Online Support First released version
   //01.00.01 20.12.2017 Siemens Industry Online Support GetStationInfo removed
   //01.00.02 27.02.2018 Siemens Industry Online Support Minor corrections
   //=============================================================================

   IF (#ioSystemHwId <> #ioSystemData.hardwareId)
   THEN
       // New IO System detected at input
       #statFirstDeviceFlag := TRUE;
       #statFirstDevice := 1;
       #statLastDevice := 1;

       #statActualConfiguredDevices := 0;
       #tempDeviceIndex := 1;

       #statError := FALSE;
       #statStatus := #STATUS_EXECUTION_FINISHED;
       #statStatusID := 0;
       #ioSystemData.error := FALSE;
       #ioSystemData.hardwareId := #ioSystemHwId;

       // Find out the number of the assigned IO system
       #tempRetValGeo := LOG2GEO(LADDR := #ioSystemHwId,
                                 GEOADDR := #statGeoAddr);
       // Set IO system ID
       #ioSystemData.number := #statGeoAddr.IOSYSTEM;

       // Initialize the structure for system function GEO2LOG
       #statGeoAddr.HWTYPE := #DEVICE_SLAVE;   // Hardware type 2: IO device

       // Predefine the type OF IO system. Either Profinet IO or Profibus DP
       IF (#statGeoAddr.AREA = #IO_SYSTEM_AREA)     // Area ID 1: PROFINET IO
       THEN
           #statMaxDevices := "USERDIAG_DEVICES_PER_IO_SYSTEM_UPPER_LIM";
       ELSIF (#statGeoAddr.AREA = #DP_SYSTEM_AREA) // Area ID 2: Profibus DP
       THEN
           IF ("USERDIAG_DEVICES_PER_IO_SYSTEM_UPPER_LIM" > #MAX_SLAVES_DP)
           THEN
               #statMaxDevices := #MAX_SLAVES_DP;
           ELSE
               #statMaxDevices := "USERDIAG_DEVICES_PER_IO_SYSTEM_UPPER_LIM";
           END_IF;
       ELSE
           #statMaxDevices := "USERDIAG_DEVICES_PER_IO_SYSTEM_UPPER_LIM";
       END_IF;

       // Set all other devices to not configured
       FOR #tempIndex := 1 TO "USERDIAG_DEVICES_PER_IO_SYSTEM_UPPER_LIM" DO
           #ioSystemData.devices[#tempIndex] := #tempDeviceInit;
       END_FOR;

       //=============================================================================
       // CONFIGURED DEVICES
       //=============================================================================
       // Find out how much devices are configured in the IO System --> PROFINET IO
       // This number is the maximum number of devices, which will be checked in the
       // following programm
       #tempRetValDeviceStates := DeviceStates(LADDR := #ioSystemHwId,
                                               MODE := #MODE_CONFIGURED,
                                               STATE := #statConfiguredDevices);

       // Check if the block call was successful
       IF (#tempRetValDeviceStates = 0)
       THEN
           // Call ok
           ;
       ELSIF (#tempRetValDeviceStates = #ERR_HWID_NOT_EXISTENT)
           OR (#tempRetValDeviceStates = #ERR_LADDR_ADDRESS)
       THEN
           #ioSystemData.error := TRUE;
           #statStatus := INT_TO_WORD(#tempRetValDeviceStates);
           #statStatusID := #ID_DEVICE_STATES_CONFIGURED;
           #statError := TRUE;
       ELSE
           // Error handling
           #statStatus := INT_TO_WORD(#tempRetValDeviceStates);
           #statStatusID := #ID_DEVICE_STATES_CONFIGURED;
           #statError := TRUE;
       END_IF;

